(* Logix 5000 project; controller FV vendor 1 type 14 code 217 rev 31.11; software revision 31.00; part 5 of 63 *)
(* tags used below, declared in another part *)
   _1s_pulse : BOOL;
   FR_ALARM_RETURNED_STRING : STRING;
   FR_Crop_Event_Prefix : STRING;
   FR_Crop_Log_ID : DINT;
   FR_Event_Alarm_Tag : ALARM_DIGITAL;
   FR_Event_control_FIFO : CONTROL;
   FR_Event_control_FIFO_Operation_Type : CONTROL;
   FR_Event_Delay_For_Data : TIMER;
   FR_Event_Delay_For_PLC_Startup_Data : TIMER;
   FR_Event_Delay_Timer : TIMER;
   FR_Event_Delay_Timer_Off : TIMER;
   FR_Event_from_buffer : STRING;
   FR_Event_from_buffer_LogData1 : REAL;
   FR_Event_from_buffer_LogData2 : REAL;
   FR_Event_from_buffer_LogData3 : REAL;
   FR_Event_from_buffer_LogData4 : REAL;
   FR_Event_from_buffer_Operation_Type : DINT;
   FR_event_step : DINT;
   FR_Event_String_Last : STRING;
   FR_Event_Transact_Trigger_Tag : DINT;
   FR_Events_FIFO_Buffer : STRING[31];
   FR_Events_FIFO_Buffer_Operation_Type : DINT[31];
   FR_Filling_Event_Prefix : STRING;
   FR_Filling_Log_ID : DINT;
   FR_Filtrate_Event_Prefix : STRING;
   FR_Filtrate_Log_ID : DINT;
   FR_FVs26_31_Cropping_Event : STRING;
   FR_FVs26_31_Filling_Event : STRING;
   FR_FVs26_31_Filtrate_Event : STRING;
   FR_FVs26_31_Green_Beer_Event : STRING;
   FR_GreenBeer_Event_Prefix : STRING;
   FR_GreenBeer_Log_ID : DINT;
   FR_Last_LogData_For_Op : REAL[30,20];
   FR_N100 : INT[265];   // FV FILLING
   FR_N100_6_alarm : ALARM_DIGITAL;
   FR_N100_6_Alarm_Ready : BOOL;
   FR_N100_6_Delayed : DINT;
   FR_N100_6_Delayed_Timer : TIMER;
   FR_N100_6_Fault_Returned : STRING;
   FR_N100_6_SQL_Done : DINT;
   FR_N100_7_alarm : ALARM_DIGITAL;
   FR_N100_7_Alarm_Ready : BOOL;
   FR_N100_7_Delayed : DINT;
   FR_N100_7_Delayed_Timer : TIMER;
   FR_N100_7_Delayed_Timer2 : TIMER;
   FR_N100_7_Fault_Returned : STRING;
   FR_N100_7_SQL_Done : DINT;
   FR_N100_8_Delayed : DINT;
   FR_N100_8_Delayed_Timer : TIMER;
   FR_N110 : INT[265];   // GREEN BEER Green Beer Main
   FR_N110_6_alarm : ALARM_DIGITAL;
   FR_N110_6_Alarm_Ready : BOOL;
   FR_N110_6_Delayed : DINT;
   FR_N110_6_Delayed_Timer : TIMER;
   FR_N110_6_Fault_Returned : STRING;
   FR_N110_6_SQL_Done : DINT;
   FR_N110_7_alarm : ALARM_DIGITAL;
   FR_N110_7_Alarm_Ready : BOOL;
   FR_N110_7_Delayed : DINT;
   FR_N110_7_Delayed_Timer : TIMER;
   FR_N110_7_Delayed_Timer2 : TIMER;
   FR_N110_7_Fault_Returned : STRING;
   FR_N110_7_SQL_Done : DINT;
   FR_N110_8_Delayed : DINT;
   FR_N110_8_Delayed_Timer : TIMER;
   FR_N120 : INT[265];   // YEAST CROP Yeast Cropping Main
   FR_N120_6_alarm : ALARM_DIGITAL;
   FR_N120_6_Alarm_Ready : BOOL;
   FR_N120_6_Delayed : DINT;
   FR_N120_6_Delayed_Timer : TIMER;
   FR_N120_6_Fault_Returned : STRING;
   FR_N120_6_SQL_Done : DINT;
   FR_N120_7_alarm : ALARM_DIGITAL;
   FR_N120_7_Alarm_Ready : BOOL;
   FR_N120_7_Delayed : DINT;
   FR_N120_7_Delayed_Timer : TIMER;
   FR_N120_7_Delayed_Timer2 : TIMER;
   FR_N120_7_Fault_Returned : STRING;
   FR_N120_7_SQL_Done : DINT;
   FR_N120_8_Delayed : DINT;
   FR_N120_8_Delayed_Timer : TIMER;
   FR_N130 : INT[265];   // FILTRATE Filtrate Return
   FR_N130_6_alarm : ALARM_DIGITAL;
   FR_N130_6_Alarm_Ready : BOOL;
   FR_N130_6_Delayed : DINT;
   FR_N130_6_Delayed_Timer : TIMER;
   FR_N130_6_Fault_Returned : STRING;
   FR_N130_6_SQL_Done : DINT;
   FR_N130_7_alarm : ALARM_DIGITAL;
   FR_N130_7_Alarm_Ready : BOOL;
   FR_N130_7_Delayed : DINT;
   FR_N130_7_Delayed_Timer : TIMER;
   FR_N130_7_Delayed_Timer2 : TIMER;
   FR_N130_7_Fault_Returned : STRING;
   FR_N130_7_SQL_Done : DINT;
   FR_N130_8_Delayed : DINT;
   FR_N130_8_Delayed_Timer : TIMER;
   FtoF_raw_input : REAL;
   FV_B22 : INT[255];   // YSVFILL_FL YSV filling process flags
   FV_B32 : INT[255];   // PITCH_FLGS YSV pitching control flags
   FV_B42 : INT[255];   // YSVCIP_FLG
   FV_B52 : INT[255];   // WASTE_FLG
   FV_B62 : INT[255];   // RESEED FLG
   FV_B82 : INT[255];   // YSTFILL FL YST filling process flags
   FV_B86 : INT[255];   // YSTCIP FL YST CIP process flag s
   FV_N101 : INT[255];   // FV INT Fermentation control integer workspace
   FV_N139 : INT[255];   // YST1
   FV_N140 : INT[255];   // YST2
   FV_N141 : INT[255];   // YSV1 DATA
   FV_N142 : INT[255];   // YSV2 DATA
   FV_N143 : INT[255];   // YSV3 DATA
   FV_N144 : INT[255];   // YST1 DATA
   FV_N145 : INT[255];   // YST2 DATA
   FV_N20 : INT[255];   // YSVFILL<PC YSV Filling data fro m PC
   FV_N21 : INT[255];   // YSVFILL>PC YSV Filling process data to PC and contr ol regs
   FV_N30 : INT[255];   // PITCH<PC YSV Pitching data fr om PC
   FV_N31 : INT[255];   // PITCH>PC YSV Pitching data at o PC and control reg isters
   FV_N40 : INT[255];   // YSVCIP<PC
   FV_N41 : INT[255];   // YSVCIP>PC
   FV_N50 : INT[255];   // WASTE<PC
   FV_N51 : INT[255];   // WASTE>PC
   FV_N60 : INT[255];   // RESEED<PC
   FV_N61 : INT[255];   // RESEED>PC
   FV_N81 : INT[255];   // YSTFILL>PC YST filling process data to PC and contr ol regs.

        [5]   // YST filling routine alarm parameter #1
        [15]   // YST filling current YST data file pointer
        [16]   // YST filling command processor current step
   FV_N81_4_alarm : ALARM_DIGITAL;
   FV_N81_4_Alarm_Ready : BOOL;
   FV_N81_4_Delayed_Timer2 : TIMER := (PRE := 1000);
   FV_N81_4_Fault_Returned : STRING;
   FV_N81_4_SQL_Done : DINT := -1;
   FV_N84 : INT[255] := ([1] := -32768, [2] := -32768, [3] := -32768, [4] := -32768, [5] := -32768, [6] := -32768, [7] := -32768);   // YSTCIP<PC YST CIP data from PC
        [0].3   // Continue YST CIP
        [1]   // YST CIP selected YST
        [0].5   // End YST CIP
        [0].0   // Initiate YST CIP startup
        [0].15   // YST CIP cancel startup
        [0]   // YST CIP selected command
        [0].1   // Start YST CIP
        [0].4   // Abort YST CIP
        [0].2   // Stop YST CIP
   FV_N85 : INT[255] := ([0] := 1, [2] := 1, [16] := 1);   // YSTCIP>PC YST CIP process data to PC and control r egs.
        [2].3   // YST CIP continue available
        [4]   // YST CIP routine alarm register
        [9]   // YST CIP PC- displayed current step
        [1]   // YST CIP process current step
        [3]   // YST CIP process restart step
        [2].2   // YST CIP stop available
        [2].1   // YST CIP start available
        [2].4   // YST CIP abort available
        [14]   // YST CIP current YST attemperation file pointer
        [16]   // YST CIP command processor current step
        [15]   // YST CIP current YST data file pointer
        [2].0   // YST CIP initiate startup available
        [2].5   // YST CIP end available
        [0]   // YST CIP status (0:Unavailable; 1:Idle; 2:Running; 3:Stopped; 4:Faulted)
   FV_N85_4_alarm : ALARM_DIGITAL;
   FV_N85_4_Alarm_Ready : BOOL;
   FV_N85_4_Delayed_Timer2 : TIMER := (PRE := 1000);
   FV_N85_4_Fault_Returned : STRING;
   FV_N85_4_SQL_Done : DINT := -1;
   FV_N88 : INT[255] := ([1] := 99, [10] := 1, [20] := 1, [22] := 2, [23] := 10, [24] := 137, [28] := 5, [34] := 11826, [35] := 11828, [36] := 12593, [37] := 12590, [38] := 12338, [40] := -16384, [42] := 2, [43] := 10, [44] := 137, [48] := 23, [54] := 14641, [55] := 11826, [56] := 13873, [57] := 11832, [58] := 12338, [59] := 13102, [60] := 56);   // YSP COMMS Data transferred to/ from yeast press PLC
        [20].0   // Comms.to Yeast Press PLC failed flag
        [1]   // This PLC -> YSP PLC target tank no.
        [11].0   // YSP PLC -> This PLC YST1 high level probe
        [11].1   // YST PLC -> This PLC YST2 high level probe
        [10].0   // YSP PLC -> This PLC comms.handshake flag
        [0].0   // This PLC -> YSP PLC comms.handshake flag
   FV_PITCH_ACT : ALIAS FOR FV_B32[0].0;   // YSV Pitching Process Active
   FV_PITCH_AVAILABL_CMD : ALIAS FOR FV_N31[2];   // YSV Pitching Available Commands
   FV_PITCH_CUR_STEP : ALIAS FOR FV_N31[1];   // YSV Pitching Current Step
   FV_PITCH_DIALOG_AVAIL : ALIAS FOR FV_N31[2].0;   // PLC>PC YSV Pitching Startup Dialog Button Available
   FV_PITCH_PSCAN : ALIAS FOR FV_B32[0].2;   // YSV Pitching Postscan oneshot
   FV_PITCH_RES_STEP : ALIAS FOR FV_N31[3];   // YSV Pitching Restart Step
   FV_PITCH_RUN : ALIAS FOR FV_B32[0].1;   // YSVPitching Running
   FV_PITCH_SELECTED_CMD : ALIAS FOR FV_N30[0];   // YSV Pitching Selected Command
   FV_PITCH_START_SELECT : ALIAS FOR FV_N30[0].0;   // PC>PLC YSV Pitching Startup Dialog Buttlon Selected
   FV_PITCH_STATUS : ALIAS FOR FV_N31[0];   // YSV Pitching Status
   FV_PUMP1 : PlantItem := (CW := 2#0000_0000_0000_0000_0000_0000_1000_0001, CheckTime := 8, DriveBits := 1);   // PUMP1
   FV_PUMP1_RawOutput : ALIAS FOR Remote_IO:4:O.Data.13;   // FV_PUMP1 Coolant recirc.valve 1
   FV_PUMP2 : PlantItem := (CW := 2#0000_0000_0000_0000_0000_0000_1010_0001, CheckTime := 8, DriveBits := 1);   // PUMP2
   FV_PUMP2_RawOutput : ALIAS FOR Remote_IO:4:O.Data.14;   // FV_PUMP2 Coolant recirc.valve 2
   FV_PUMP3 : PlantItem := (CheckTime := 8);   // PUMP3
   FV_PUMP3_RawOutput : ALIAS FOR Remote_IO:4:O.Data.15;   // FV_PUMP3 Coolant recirc.valve 3
   FV_PV550_DPTR : ALIAS FOR FV_N101[8];   // Fermenting Room PV550 data file pointer
   FV_PX1 : PlantItem := (CW := 2#0000_0000_0000_0100_0000_0000_0000_0001, CheckTime := 12, DebounceTime := 4);   // PX1
   FV_PX1_RawInput : ALIAS FOR Remote_IO:6:I.Data.13;   // FV_PX1 Water flush proxy switch
   FV_PX2 : PlantItem := (CW := 2#0000_0000_0000_0000_0000_0000_0010_0000);   // PX2
   FV_PX2_RawInput : ALIAS FOR Remote_IO:6:I.Data.14;   // FV_PX2 CIP supply proxy switch
   FV_PX3 : PlantItem := (CW := 2#0000_0000_0000_0100_0000_0000_0010_0001);   // PX3
   FV_PX3_RawInput : ALIAS FOR Remote_IO:6:I.Data.15;   // FV_PX3 YSV1 to reseeding main proxy switch
   FV_R2V1 : PlantItem := (CW := 2#0000_0000_0000_0000_0000_0000_0001_0000, CheckTime := 15, CheckTimer := 15);   // R2V1
   FV_R2V1_ALARM : ALARM_DIGITAL;
   FV_R2V1_C : ALIAS FOR Remote_IO:7:I.Data.6;
   FV_R2V1_DR : ALIAS FOR Remote_IO:5:O.Data.10;
   FV_R2V1_O : ALIAS FOR Remote_IO:7:I.Data.2;
   FV_R2V2 : PlantItem := (CW := 2#0000_0000_0000_0000_0000_0000_1000_1011, CheckTime := 4, CheckTimer := 4, DriveBits := 4);   // R2V2
   FV_R2V2_ALARM : ALARM_DIGITAL;
   FV_R2V2_C : ALIAS FOR Remote_IO:7:I.Data.7;
   FV_R2V2_DR : ALIAS FOR Remote_IO:5:O.Data.11;
   FV_R2V2_O : ALIAS FOR Remote_IO:7:I.Data.3;
   FV_R6 : CONTROL[5] := ([1].LEN := 3, [2].LEN := 3, [2].UL := 1, [3].LEN := 3);
   FV_RESEED_ACT : ALIAS FOR FV_B62[0].0;   // YSV Reseeding Process Active
   FV_RESEED_AV1 : ALIAS FOR FV_B62[1];
   FV_RESEED_AV2 : ALIAS FOR FV_B62[2];
   FV_RESEED_AV3 : ALIAS FOR FV_B62[3];
   FV_RESEED_AV4 : ALIAS FOR FV_B62[4];
   FV_RESEED_AV5 : ALIAS FOR FV_B62[5];
   FV_RESEED_AVAILABL_CMD : ALIAS FOR FV_N61[2];   // YSV Reseeding Available Commands
   FV_RESEED_CUR_STEP : ALIAS FOR FV_N61[1];   // YSV Reseeding Current Step
   FV_RESEED_DIALOG_AVAIL : ALIAS FOR FV_N61[2].0;   // PLC>PC YSV Reseeding Startup Dialog Button Available
   FV_RESEED_END : ALIAS FOR FV_B62[0].8;   // YSV Reseeding End Process Selected
   FV_RESEED_PSCAN : ALIAS FOR FV_B62[0].2;   // YSV Reseeding Postscan oneshot
   FV_RESEED_RES_STEP : ALIAS FOR FV_N61[3];   // YSV Reseeding Restart Step
   FV_RESEED_RUN : ALIAS FOR FV_B62[0].1;   // YSV Reseeding Running
   FV_RESEED_SELECTED_CMD : ALIAS FOR FV_N60[0];   // YSV Reseeding Selected Command
   FV_RESEED_START_SELECT : ALIAS FOR FV_N60[0].0;   // PC>PLC YSV Reseeding Startup Dialog Buttlon Selected
   FV_RESEED_STATUS : ALIAS FOR FV_N61[0];   // YSV Reseeding Status
   FV_RSLN_CLEAN : ALIAS FOR FV_B62[1].0;   // Reseeding line clean flag
   FV_SFile : INT[255] := ([4] := 19904, [13] := 3, [37] := 2020, [38] := 7, [39] := 31, [40] := 13, [41] := 9, [42] := 50);   // SLC Equivalent System File, So Original Code Can Remain
        [1].15   // First Scan Flag
        [37]   // Clock Calendar Year
        [41]   // Clock Calendar Minutes
        [53]   // Calendar Day 1 = Monday
        [40]   // Clock Calendar Hours
        [42]   // Clock Calendar Minute
   FV_SOV1 : PlantItem := (CheckTime := 8);   // SOV1
   FV_SOV1_RawOutput : ALIAS FOR Remote_IO:5:O.Data.6;   // FV_SOV1 Air supply to reseed pump
   FV_SOV2 : PlantItem := (CheckTime := 8);   // SOV2
   FV_SOV2_RawOutput : ALIAS FOR Remote_IO:5:O.Data.7;   // FV_SOV2 Air supply to reseed pump
   FV_T102 : TIMER[20] := ([0].PRE := 360000, [0].ACC := 298181, [0].EN := 1, [0].TT := 1);
   FV_T16 : TIMER[10] := ([0].PRE := 8000, [0].ACC := 3002, [0].EN := 1, [0].TT := 1);
   FV_T212 : TIMER[5] := ([0].PRE := 3000, [0].EN := 1, [0].DN := 1, [1].PRE := 3000, [1].EN := 1, [1].DN := 1, [2].PRE := 3000, [2].ACC := 3000);
   FV_T23 : TIMER[10] := ([0].PRE := 300000);
   FV_T33 : TIMER[10] := ([0].PRE := 300000, [1].PRE := 60000, [2].PRE := 10000);
   FV_T4 : TIMER[10] := ([0].PRE := 2000, [1].PRE := 300000, [2].PRE := 2500, [2].ACC := 50, [2].EN := 1, [2].TT := 1, [3].PRE := 300000, [3].ACC := 300001, [3].EN := 1, [3].DN := 1, [4].PRE := 3300000, [4].ACC := 2309456, [4].EN := 1, [4].TT := 1, [5].PRE := 3600000, [6].PRE := 60000, [8].PRE := 10000, [9].PRE := 10000);
   FV_T43 : TIMER[10] := ([0].PRE := 300000);
   FV_T53 : TIMER[10] := ([0].PRE := 300000, [2].PRE := 10000);
   FV_T63 : TIMER[20] := ([0].PRE := 60000, [3].PRE := 120000, [3].ACC := 82385, [4].PRE := 13000, [5].PRE := 16000, [6].PRE := 30000, [7].PRE := 4000, [8].PRE := 4000);
   FV_T73 : TIMER[10] := ([0].PRE := 300000, [1].PRE := 30000, [2].PRE := 20000);
   FV_T83 : TIMER[5] := ([0].PRE := 300000);
   FV_T87 : TIMER[2] := ([0].PRE := 300000);
   FV_T89 : TIMER[5] := ([0].PRE := 3000, [0].ACC := 1745, [0].EN := 1, [0].TT := 1, [1].PRE := 10000, [2].PRE := 10000, [2].ACC := 10001, [2].EN := 1, [2].DN := 1);
   FV_to_data_file : DINT;
   FV_to_data_offset : DINT;
   FV_TTX_YS_001_AI : PlantItem := (CW := 2#0000_0000_0000_0000_1100_0000_0000_0000, CheckTime := 10, CheckTimer := 10, Scaled := 18.41875, RawInput := 6947.0);   // TTX_YS_001
   FV_TTX_YS_001_AI_RawInput : ALIAS FOR Remote_IO:8:I.Ch00Data;   // Real Analog Input , Do Not Use In Code
   FV_TTX_YS_002_AI : PlantItem := (CW := 2#0000_0000_0000_0000_1000_0000_0000_0000, CheckTime := 10, CheckTimer := 10, Scaled := 9.6625, RawInput := 5546.0);   // TTX_YS_002
   FV_TTX_YS_002_AI_RawInput : ALIAS FOR Remote_IO:8:I.Ch01Data;   // Real Analog Input , Do Not Use In Code
   FV_value_to_set : INT;
   FV_WASTE_ACT : ALIAS FOR FV_B52[0].0;   // YSV To Waste Process Active
   FV_WASTE_AVAILABL_CMD : ALIAS FOR FV_N51[2];   // YSV To Waste Available Commands
   FV_WASTE_CUR_STEP : ALIAS FOR FV_N51[1];   // YSV To Waste Current Step
   FV_WASTE_DIALOG_AVAIL : ALIAS FOR FV_N51[2].0;   // PLC>PC YSV To Waste Startup Dialog Button Available
   FV_WASTE_PSCAN : ALIAS FOR FV_B52[0].2;   // YSV To Waste Postscan oneshot
   FV_WASTE_RES_STEP : ALIAS FOR FV_N51[3];   // YSV To Waste Restart Step
   FV_WASTE_RUN : ALIAS FOR FV_B52[0].1;   // YSV To Waste Running
   FV_WASTE_SELECTED_CMD : ALIAS FOR FV_N50[0];   // YSV To Waste Selected Command
   FV_WASTE_START_SELECT : ALIAS FOR FV_N50[0].0;   // PC>PLC YSV To Waste Startup Dialog Buttlon Selected
   FV_WASTE_STATUS : ALIAS FOR FV_N51[0];   // YSV To Waste Status
   FV_word_offset : INT;
   FV_WYT1R : PlantItem := (CW := 2#0000_0000_0000_0000_0000_1100_0000_0000, CheckTime := 8, CheckTimer := 8);   // WYT1R
   FV_WYT1R_ALARM : ALARM_DIGITAL;
   FV_WYT1R_D : ALIAS FOR Remote_IO:5:O.Data.14;
   FV_WYT1R_R : ALIAS FOR Remote_IO:7:I.Data.20;
   FV_WYT2R : PlantItem := (CW := 2#0000_0000_0000_0000_0000_1100_1000_1011, CheckTime := 8, CheckTimer := 8, DriveBits := 1);   // WYT2R
   FV_WYT2R_ALARM : ALARM_DIGITAL;
   FV_WYT2R_D : ALIAS FOR Remote_IO:5:O.Data.15;
   FV_WYT2R_R : ALIAS FOR Remote_IO:7:I.Data.21;
   FV_WYTR1 : PlantItem := (CW := 2#0000_0000_0000_0000_0000_0000_0001_0000, CheckTime := 10, CheckTimer := 10);   // WYTR1
   FV_WYTR1_ALARM : ALARM_DIGITAL;
   FV_WYTR1_C : ALIAS FOR Remote_IO:7:I.Data.4;
   FV_WYTR1_DR : ALIAS FOR Remote_IO:5:O.Data.8;
   FV_WYTR1_O : ALIAS FOR Remote_IO:7:I.Data.0;
   FV_WYTR2 : PlantItem := (CW := 2#0000_0000_0000_0000_0000_0000_0001_0000, CheckTime := 4, CheckTimer := 4);   // WYTR2
   FV_WYTR2_ALARM : ALARM_DIGITAL;
   FV_WYTR2_C : ALIAS FOR Remote_IO:7:I.Data.5;
   FV_WYTR2_DR : ALIAS FOR Remote_IO:5:O.Data.9;
   FV_WYTR2_O : ALIAS FOR Remote_IO:7:I.Data.1;
   FV_Yeast_Press_Blunger_Comms : MESSAGE;
        MessageParameters(ServiceCode := 16#0fa2, LocalElement := FV_N88[10], ...)
   FV_YSPC_FAIL : ALIAS FOR FV_N88[20].0;   // Comms.to Yeast Press PLC failed flag
   FV_YST01_LTX501_Fill_Lvl_OK : TIMER := (PRE := 1000);
   FV_YST02_LTX501_Fill_Lvl_OK : TIMER := (PRE := 1000);
   FV_YST1_FV : ALIAS FOR FV_N139[0];   // YST1 attemperation control data
   FV_YST1_HL_SP : DINT := 145;
   FV_YST1_STATUS : ALIAS FOR FV_N144[0];   // YST1 current operation
   FV_YST2_FV : ALIAS FOR FV_N140[0];   // YST2 attemperation control data
   FV_YST2_HL_SP : DINT := 145;
   FV_YST2_STATUS : ALIAS FOR FV_N145[0];   // YST2 current operation
   FV_YSTCIP_ACT : ALIAS FOR FV_B86[0].0;   // YST CIP process active
   FV_YSTCIP_Log_ID : DINT := 10;
   FV_YSTCIP_RESTART : ALIAS FOR FV_N85[3];   // YST CIP process restart step
   FV_YSTCIP_RUN : ALIAS FOR FV_B86[0].1;   // YST CIP running
   FV_YSTCIP_STATUS : ALIAS FOR FV_N85[0];   // YST CIP status (0:Unavailable; 1:Idle; 2:Running; 3:Stopped; 4:Faulted)
   FV_YSTCIP_STEP : ALIAS FOR FV_N85[1];   // YST CIP process current step
   FV_YSTFILL_ACT : ALIAS FOR FV_B82[0].0;   // YST filling process active
   FV_YSTFILL_Log_ID : DINT := 3;
   FV_YSTFILL_PSCAN : ALIAS FOR FV_B82[0].2;   // YST filling postscan oneshot
   FV_YSTFILL_RESTART : ALIAS FOR FV_N81[3];   // YST filling restart step
   FV_YSTFILL_RUN : ALIAS FOR FV_B82[0].1;   // YST filling process running
   FV_YSTFILL_STATUS : ALIAS FOR FV_N81[0];   // YST filling status (0:Unavailable; 1:Idle; 2:Running; 3:Stopped; 4:Faulted)
   FV_YSTFILL_STEP : ALIAS FOR FV_N81[1];   // YST filling current step
   FV_YSTs_CIP_Vessel_Event : STRING;
   FV_YSTs_CIP_Vessel_Event_Prefix : STRING := 'YST 1 ';
   FV_YSTs_Filling_Event : STRING;
   FV_YSTs_Filling_Event_Prefix : STRING := 'YST 1 ';
   FV_YSV1_RSR_MODE : ALIAS FOR FV_N141[3];   // YSV1 Rouser Mode 0=Auto 1 = Manual On 2 = Manual Off
   FV_YSV1_STATUS : ALIAS FOR FV_N141[0];   // YSV1 Current Operation
   FV_YSV1_TTX01_AI : PlantItem := (CW := 2#0000_0000_0000_0000_1000_0000_0000_0000, CheckTime := 10, CheckTimer := 10, Scaled := 4.640625, RawInput := 8685.0);   // YSV1_TTX01
   FV_YSV1_TTX01_AI_RawInput : ALIAS FOR Remote_IO:13:I.Ch1Data;   // Real Analog Input , Do Not Use In Code
   FV_YSV1_WEIGHT : ALIAS FOR FV_N141[2];   // YSV1 current weight kg*10
   FV_YSV1_WTX01_AI : PlantItem := (CW := 2#0000_0000_0000_0000_1000_0000_0000_0000, CheckTime := 10, CheckTimer := 10, Scaled := 51.7575, RawInput := 5648.0);   // YSV1_WTX01
   FV_YSV1_WTX01_AI_RawInput : ALIAS FOR Remote_IO:13:I.Ch6Data;   // Real Analog Input , Do Not Use In Code
   FV_YSV1CV : PlantItem := (CW := 2#0000_0000_0000_0000_0000_0000_0100_0000, CheckTime := 8);   // YSV1CV
   FV_YSV1CV_RawOutput : ALIAS FOR Remote_IO:5:O.Data.12;   // FV_YSV1CV
   FV_YSV1J : PlantItem := (CW := 2#0000_0000_0000_0000_0000_0000_1000_0001, CheckTime := 8, DriveBits := 1);   // YSV1J
   FV_YSV1J_RawOutput : ALIAS FOR Remote_IO:4:O.Data.9;   // FV_YSV1J YSV 1 cooling valve
   FV_YSV1R : PlantItem := (CW := 2#0000_0000_0000_0000_0000_1100_0000_0000, CheckTime := 8, CheckTimer := 8);   // YSV1R
   FV_YSV1R_ALARM : ALARM_DIGITAL;
   FV_YSV1R_D : ALIAS FOR Remote_IO:4:O.Data.10;   // YSV 1 rouser
   FV_YSV1R_R : ALIAS FOR Remote_IO:6:I.Data.12;   // YSV 1 Rouser running f/b
   FV_YSV2_STATUS : ALIAS FOR FV_N142[0];   // YSV2 Current Operation
   FV_YSV2_TTX01_AI : PlantItem := (CW := 2#0000_0000_0000_0000_1000_0000_0000_0000, CheckTime := 10, CheckTimer := 10, Scaled := 3.1531248, RawInput := 8209.0);   // YSV2_TTX01
   FV_YSV2_TTX01_AI_RawInput : ALIAS FOR Remote_IO:13:I.Ch2Data;   // Real Analog Input , Do Not Use In Code
   FV_YSV2_WEIGHT : ALIAS FOR FV_N142[2];   // YSV2 current weight kg*10
   FV_YSV2_WTX01_AI : PlantItem := (CW := 2#0000_0000_0000_0000_1000_0000_0000_0000, CheckTime := 10, CheckTimer := 10, Scaled := 155.11562, RawInput := 11091.0);   // YSV2_WTX01
   FV_YSV2_WTX01_AI_RawInput : ALIAS FOR Remote_IO:13:I.Ch5Data;   // Real Analog Input , Do Not Use In Code
   FV_YSV2CV : PlantItem := (CW := 2#0000_0000_0000_0000_0000_0000_1000_0001, CheckTime := 8, DriveBits := 1);   // YSV2CV
   FV_YSV2CV_RawOutput : ALIAS FOR Remote_IO:5:O.Data.13;   // FV_YSV2CV
   FV_YSV2J : PlantItem := (CW := 2#0000_0000_0000_0000_0000_0000_1000_0001, CheckTime := 8, DriveBits := 1);   // YSV2J
   FV_YSV2J_RawOutput : ALIAS FOR Remote_IO:4:O.Data.11;   // FV_YSV2J YSV 2 cooling valve
   FV_YSV2O : PlantItem := (CheckTime := 8);   // YSV2O
   FV_YSV2O_RawOutput : ALIAS FOR Remote_IO:4:O.Data.4;   // FV_YSV2O YSV 2 outlet valve
   FV_YSV2R : PlantItem := (CheckTime := 8);   // YSV2R
   FV_YSV2R_RawOutput : ALIAS FOR Remote_IO:4:O.Data.12;   // FV_YSV2R YSV 2 rouser
   FV_YSV3_STATUS : ALIAS FOR FV_N143[0];   // YSV3 Current Operation
   FV_YSV3_TTX01_AI : PlantItem := (CW := 2#0000_0000_0000_0000_1000_0000_0000_0000, CheckTime := 10, CheckTimer := 10, Scaled := 21.153126, RawInput := 13969.0);   // YSV3_TTX01
   FV_YSV3_TTX01_AI_RawInput : ALIAS FOR Remote_IO:13:I.Ch3Data;   // Real Analog Input , Do Not Use In Code
   FV_YSV3_WEIGHT : ALIAS FOR FV_N143[2];   // YSV3 current weight kg*10
   FV_YSV3_WTX01_AI : PlantItem := (CW := 2#0000_0000_0000_0000_1000_0000_0000_0000, CheckTime := 10, CheckTimer := 10, Scaled := 0.0625, RawInput := 4002.0);   // YSV3_WTX01
   FV_YSV3_WTX01_AI_RawInput : ALIAS FOR Remote_IO:13:I.Ch4Data;   // Real Analog Input , Do Not Use In Code
   FV_YSV3J : PlantItem := (CheckTime := 8);   // YSV3J
   FV_YSV3J_RawOutput : ALIAS FOR Remote_IO:4:O.Data.7;   // FV_YSV3J YSV 3 cooling valve
   FV_YSV3O : PlantItem := (CheckTime := 8);   // YSV3O
   FV_YSV3O_RawOutput : ALIAS FOR Remote_IO:4:O.Data.6;   // FV_YSV3O YSV 3 outlet valve
   FV_YSV3R : PlantItem := (CheckTime := 8);   // YSV3R
   FV_YSV3R_RawOutput : ALIAS FOR Remote_IO:4:O.Data.8;   // FV_YSV3R YSV 3 rouser
   FV_YSVCIP_ACT : ALIAS FOR FV_B42[0].0;   // YSV CIP Process Active
   FV_YSVCIP_AVAILABL_CMD : ALIAS FOR FV_N41[2];   // YSV CIP Available Commands
   FV_YSVCIP_CUR_STEP : ALIAS FOR FV_N41[1];   // YSV CIP Current Step
   FV_YSVCIP_DIALOG_AVAIL : ALIAS FOR FV_N41[2].0;   // PLC>PC YSV CIP Startup Dialog Button Available
   FV_YSVCIP_END : ALIAS FOR FV_B42[0].8;   // YSV CIP End Process Selected
   FV_YSVCIP_PSCAN : ALIAS FOR FV_B42[0].2;   // YSV CIP Postscan oneshot
   FV_YSVCIP_RES_STEP : ALIAS FOR FV_N41[3];   // YSV CIP Restart Step
   FV_YSVCIP_RUN : ALIAS FOR FV_B42[0].1;   // YSV CIP Running
   FV_YSVCIP_SELECTED_CMD : ALIAS FOR FV_N40[0];   // YSV CIP Selected Command
   FV_YSVCIP_START_SELECT : ALIAS FOR FV_N40[0].0;   // PC>PLC YSV CIP Startup Dialog Buttlon Selected
   FV_YSVCIP_STATUS : ALIAS FOR FV_N41[0];   // YSV CIP Status
   FV_YSVCIPLINE_Log_ID : DINT := 7;
   FV_YSVCIPVESSEL_Log_ID : DINT := 6;
   FV_YSVFILL_ACT : ALIAS FOR FV_B22[0].0;   // YSV Filling Process Active
   FV_YSVFILL_AVAILABL_CMD : ALIAS FOR FV_N21[2];   // YSV Filling Available Commands
   FV_YSVFILL_CUR_STEP : ALIAS FOR FV_N21[1];   // YSV Filling Current Step
   FV_YSVFILL_DIALOG_AVAIL : ALIAS FOR FV_N21[2].0;   // PLC>PC YSV Filling Startup Dialog Button Available
   FV_YSVFILL_END : ALIAS FOR FV_B22[0].8;   // YSV Filling End Process Selected
   FV_YSVFILL_Log_ID : DINT := 4;
   FV_YSVFILL_PSCAN : ALIAS FOR FV_B22[0].2;   // YSV Filling Postscan oneshot
   FV_YSVFILL_RES_STEP : ALIAS FOR FV_N21[3];   // YSV Filling Restart Step
   FV_YSVFILL_RUN : ALIAS FOR FV_B22[0].1;   // YSV Filling Running
   FV_YSVFILL_SELECTED_CMD : ALIAS FOR FV_N20[0];   // YSV Filling Selected Command
   FV_YSVFILL_START_SELECT : ALIAS FOR FV_N20[0].0;   // PC>PLC YSV Filling Startup Dialog Buttlon Selected
   FV_YSVFILL_STATUS : ALIAS FOR FV_N21[0];   // YSV Filling Status
   FV_YSVPITCH_Log_ID : DINT := 5;
   FV_YSVPitching_AmountAtEnd : REAL := 155.68437;
   FV_YSVRESEED_Log_ID : DINT := 9;
   FV_YSVs_CIP_Line_Event : STRING;
   FV_YSVs_CIP_Line_Event_prefix : STRING;
   FV_YSVs_CIP_vessel_Event : STRING;
   FV_YSVs_CIP_vessel_Event_Prefix : STRING := 'YSV 2 ';
   FV_YSVs_Filling_Event : STRING;
   FV_YSVs_Filling_Event_Prefix : STRING := 'YSV 2 ';
   FV_YSVs_Pitching_Event : STRING;
   FV_YSVs_Pitching_Event_Prefix : STRING := 'YSV 2 ';
   FV_YSVs_reseeding_event : STRING;
   FV_YSVs_reseeding_event_prefix : STRING := 'YSV 1 ';
   FV_YSVs_to_waste_event : STRING;
   FV_YSVs_to_waste_event_prefix : STRING := 'YSV 2 ';
   FV_YSVTOWASTE_Log_ID : DINT := 8;
   FV_YSVWaste_AmountAtEnd : REAL := 0.56874996;
   go_test_operation_temp : BOOL;
   indirect_bit_temp : INT := 7;
   Item_Faults_Are_Latched : BOOL;
   Item_Simulation_Flag : BOOL;
   ItoF_raw_input : INT := 5648;
   Mike_141019 : BOOL := 1;
   MV_Read_YST : MESSAGE;
        MessageParameters(ServiceCode := 16#004c, LocalElement := MV_YST_Levels[0], ...)
   MV_Read_YST_TMR : TIMER := (PRE := 500, ACC := 485, EN := 1, TT := 1);
   MV_YST_Levels : REAL[2] := ([0] := 0.028125001, [1] := 79.640625);
        [0]   // YST1 Level
        [1]   // YST2 Level
   One_Minute_One_Scan : BOOL;
   One_Minute_One_Scan_Timer : TIMER := (PRE := 60000, ACC := 51773, EN := 1, TT := 1);
   One_Second_1_scan : BOOL;
   One_Second_One_Scan : ALIAS FOR One_Second_1_scan;
   One_Second_Toggle : BOOL := 1;
   overrange_RIO_analog_value : REAL;
   Pitching_transaction_locked_timer : TIMER := (PRE := 10000);
   Pitching_transaction_log : DINT;
   Pitching_transaction_log_delay : DINT;
   Pitching_transaction_log_Done : DINT := -1;
   Pitching_transaction_log_timer : TIMER := (PRE := 10000);
   rack_simulation_flag : BOOL;
   Reseeding_transaction_locked_timer : TIMER := (PRE := 10000);
   Reseeding_transaction_log : DINT;
   Reseeding_transaction_log_delay : DINT;
   Reseeding_transaction_log_Done : DINT := -1;
   Reseeding_transaction_log_timer : TIMER := (PRE := 10000);
   reset_msg_interval : BOOL;
   Scada_Pump_Fault_No : DINT := 20001;
   Scada_Pump_H_Fault_No : DINT;
   Scada_Pump_T_Fault_No : DINT;
   Scada_Valve_Fault_No : DINT := 10001;
   scada_watchdog : DINT := 15;
   scada_watchdog_tmr : TIMER := (PRE := 1000);
   scada_watchdog_tmr_off : TIMER := (PRE := 1000, ACC := 242, EN := 1, TT := 1);
   scale_analog_int : DINT := 12000;
   scale_analog_result : REAL := 1142.0016;
   scale_eu_max : REAL := 502.5;
   scale_eu_max_int : DINT := 300;
   scale_eu_min : REAL;
   scale_eu_min_int : DINT := 200;
   scale_raw_input : REAL := 11091.0;
   scale_raw_max : REAL := 20000.0;
   scale_raw_max_int : DINT := 120;
   scale_raw_min : REAL := 4000.0;
   scale_raw_min_int : DINT;
   scale_routine_active : BOOL := 1;
   scale_temp : REAL := 0.03140625;
   TempChecktime : DINT := 32;
   template_analog_input : PlantItem;
   template_analog_input_RawInput : REAL;
   template_analog_output : PlantItem;
   template_analog_output_RawOutput : REAL;
   template_boolean : BOOL;
   template_input : PlantItem;
   template_input_RawInput : ALIAS FOR template_boolean;
   template_output : PlantItem;
   template_output_RawOutput : ALIAS FOR template_boolean;   // P04CHILLRUN Chiller Run Signal
   template_pump : PlantItem;
   template_pump_D : ALIAS FOR template_boolean;   // auto start vacuum pump 1
   template_pump_H : ALIAS FOR template_boolean;   // vacuum pump 1 auto avail
   template_pump_ISOL : ALIAS FOR template_boolean;
   template_pump_R : ALIAS FOR template_boolean;   // vacuum pump 1 running
   template_valve : PlantItem;
   template_valve_C : ALIAS FOR template_boolean;   // skim manifold to ycv2 drain valve closed
   template_valve_DR : ALIAS FOR template_boolean;   // drive open skim manifold to ycv2 drain valve
   template_valve_O : ALIAS FOR template_boolean;   // skim manifold to ycv2 drain valve opened
   tempv : DINT;
   Test_Cropping_done : BOOL := 1;
   underrange_RIO_analog_value : REAL;
   Unused_Healthy_Feedback : BOOL := 1;
   Unused_NotTripped_Feedback : BOOL := 1;
   YP_ALARM_ACCEPT : ALIAS FOR YP_B103[1].2;
   YP_ALARM_ACCEPT_OS_FLAG : ALIAS FOR YP_B103[1].0;
   YP_AV1 : PlantItem := (CW := 2#0000_0000_0000_0000_0000_0000_0001_0000, CheckTime := 15, CheckTimer := 15);   // AV1
   YP_AV10_MANUAL : ALIAS FOR YP_N50[9];
   YP_AV10_REQUIRED : ALIAS FOR YP_B30[0].14;   // BLUNGER TRANSFER PUMP
   YP_AV1_ALARM : ALARM_DIGITAL;
   YP_AV1_CLOSE_FAULT : ALIAS FOR YP_B92[0].1;
   YP_AV1_CLOSE_FLT_TIMER : ALIAS FOR YP_T20[1];
   YP_AV1_DR : ALIAS FOR RIO_Rack_3:3:O.Data.3;
   YP_AV1_MANUAL : ALIAS FOR YP_N50[0];
   YP_AV1_O : ALIAS FOR RIO_Rack_3:1:I.Data.0;
   YP_AV1_OPEN_FAULT : ALIAS FOR YP_B92[0].0;
   YP_AV1_OPEN_FLT_TIMER : ALIAS FOR YP_T20[0];
   YP_AV1_REQUIRED : ALIAS FOR YP_B30[0].3;
   YP_AV2 : PlantItem := (CW := 2#0000_0000_0000_0000_0000_0001_0001_0000, CheckTime := 15, CheckTimer := 15);   // AV2
   YP_AV2_ALARM : ALARM_DIGITAL;
   YP_AV2_CLOSE_FAULT : ALIAS FOR YP_B92[0].3;
   YP_AV2_CLOSE_FLT_TIMER : ALIAS FOR YP_T20[3];
   YP_AV2_DR : ALIAS FOR RIO_Rack_3:3:O.Data.5;
   YP_AV2_MANUAL : ALIAS FOR YP_N50[1];
   YP_AV2_O : ALIAS FOR RIO_Rack_3:1:I.Data.2;
   YP_AV2_OPEN_FAULT : ALIAS FOR YP_B92[0].2;
   YP_AV2_OPEN_FLAG : ALIAS FOR YP_B3[0].2;
   YP_AV2_OPEN_FLT_TIMER : ALIAS FOR YP_T20[2];
   YP_AV2_REQUIRED : ALIAS FOR YP_B30[0].5;
   YP_AV3 : PlantItem := (CW := 2#0000_0000_0000_0000_0000_0000_0001_0000, CheckTime := 15, CheckTimer := 15);   // AV3
   YP_AV3_ALARM : ALARM_DIGITAL;
   YP_AV3_CLOSE_FAULT : ALIAS FOR YP_B92[0].5;
   YP_AV3_CLOSE_FLT_TIMER : ALIAS FOR YP_T20[5];
   YP_AV3_DR : ALIAS FOR RIO_Rack_3:3:O.Data.6;
   YP_AV3_MANUAL : ALIAS FOR YP_N50[2];
   YP_AV3_O : ALIAS FOR RIO_Rack_3:1:I.Data.4;
   YP_AV3_OPEN_FAULT : ALIAS FOR YP_B92[0].4;
   YP_AV3_OPEN_FLAG : ALIAS FOR YP_B3[0].4;
   YP_AV3_OPEN_FLT_TIMER : ALIAS FOR YP_T20[4];
   YP_AV3_REQUIRED : ALIAS FOR YP_B30[0].6;
   YP_AV4 : PlantItem := (CW := 2#0000_0000_0000_0000_0000_0000_0001_0000, CheckTime := 15, CheckTimer := 15);   // AV4
   YP_AV4_ALARM : ALARM_DIGITAL;
   YP_AV4_CLOSE_FAULT : ALIAS FOR YP_B92[0].7;
   YP_AV4_CLOSE_FLT_TIMER : ALIAS FOR YP_T20[7];
   YP_AV4_DR : ALIAS FOR RIO_Rack_3:3:O.Data.7;
   YP_AV4_MANUAL : ALIAS FOR YP_N50[3];
   YP_AV4_O : ALIAS FOR RIO_Rack_3:1:I.Data.6;
   YP_AV4_OPEN_FAULT : ALIAS FOR YP_B92[0].6;
   YP_AV4_OPEN_FLAG : ALIAS FOR YP_B3[0].6;
   YP_AV4_OPEN_FLT_TIMER : ALIAS FOR YP_T20[6];
   YP_AV4_REQUIRED : ALIAS FOR YP_B30[0].7;
   YP_AV5 : PlantItem := (CW := 2#0000_0000_0000_0000_0000_0000_0001_0000, CheckTime := 15, CheckTimer := 15);   // AV5
   YP_AV5_ALARM : ALARM_DIGITAL;
   YP_AV5_CLOSE_FLT_TIMER : ALIAS FOR YP_T20[9];
   YP_AV5_CLSOE_FAULT : ALIAS FOR YP_B92[0].9;
   YP_AV5_DR : ALIAS FOR RIO_Rack_3:3:O.Data.8;
   YP_AV5_O : ALIAS FOR RIO_Rack_3:1:I.Data.8;
   YP_AV5_OPEN_FAULT : ALIAS FOR YP_B92[0].8;
   YP_AV5_OPEN_FLAG : ALIAS FOR YP_B3[0].8;
   YP_AV5_OPEN_FLT_TIMER : ALIAS FOR YP_T20[8];
   YP_AV5_REQUIRED : ALIAS FOR YP_B30[0].8;
   YP_AV6 : PlantItem := (CW := 2#0000_0000_0000_0000_0000_0000_0001_0000, CheckTime := 15, CheckTimer := 15);   // AV6
   YP_AV6_ALARM : ALARM_DIGITAL;
   YP_AV6_CLOSE_FAULT : ALIAS FOR YP_B92[0].11;
   YP_AV6_CLOSE_FLT_TIMER : ALIAS FOR YP_T20[11];
   YP_AV6_DR : ALIAS FOR RIO_Rack_3:3:O.Data.9;
   YP_AV6_MANUAL : ALIAS FOR YP_N50[5];
   YP_AV6_O : ALIAS FOR RIO_Rack_3:1:I.Data.10;
   YP_AV6_OPEN_FAULT : ALIAS FOR YP_B92[0].10;
   YP_AV6_OPEN_FLAG : ALIAS FOR YP_B3[0].10;
   YP_AV6_OPEN_FLT_TIMER : ALIAS FOR YP_T20[10];
   YP_AV6_RQUIRED : ALIAS FOR YP_B30[0].9;
   YP_AV7 : PlantItem := (CW := 2#0000_0000_0000_0000_0000_0000_0001_0000, CheckTime := 15, CheckTimer := 15);   // AV7
   YP_AV7_ALARM : ALARM_DIGITAL;
   YP_AV7_CLOSE_FAULT : ALIAS FOR YP_B92[0].13;
   YP_AV7_CLOSE_FLT_TIMER : ALIAS FOR YP_T20[13];
   YP_AV7_DR : ALIAS FOR RIO_Rack_3:3:O.Data.10;
   YP_AV7_MANUAL : ALIAS FOR YP_N50[6];
   YP_AV7_O : ALIAS FOR RIO_Rack_3:1:I.Data.12;
   YP_AV7_OPEN_FAULT : ALIAS FOR YP_B92[0].12;
   YP_AV7_OPEN_FLAG : ALIAS FOR YP_B3[0].12;
   YP_AV7_OPEN_FLT_TIMER : ALIAS FOR YP_T20[12];
   YP_AV7_REQUIRED : ALIAS FOR YP_B30[0].10;
   YP_AV8 : PlantItem := (CW := 2#0000_0000_0000_0000_0000_0000_0001_0000, CheckTime := 15, CheckTimer := 15);   // AV8
   YP_AV8_ALARM : ALARM_DIGITAL;
   YP_AV8_CLOSE_FAULT : ALIAS FOR YP_B92[0].15;
   YP_AV8_CLOSE_FLT_TIMER : ALIAS FOR YP_T20[15];
   YP_AV8_DR : ALIAS FOR RIO_Rack_3:3:O.Data.11;
   YP_AV8_MANUAL : ALIAS FOR YP_N50[7];
   YP_AV8_O : ALIAS FOR RIO_Rack_3:1:I.Data.14;
   YP_AV8_OPEN_FAULT : ALIAS FOR YP_B92[0].14;
   YP_AV8_OPEN_FLAG : ALIAS FOR YP_B3[0].14;
   YP_AV8_OPEN_FLT_TIMER : ALIAS FOR YP_T20[14];
   YP_AV8_REQUIRED : ALIAS FOR YP_B30[0].11;
   YP_AV9_MANUAL : ALIAS FOR YP_N50[8];
   YP_B103 : INT[15] := ([0] := 1);   // Original N File From SLC, No Description Available
        [0].0   // Yeast Press CIP Heartbeat Fault
        [2].2   // Channel 1 CIP Active
        [2].3   // Channel 2 CIP Active
        [3].0   // START BLUNGER WATER FILL FROM PV
        [3].1   // STOP BLUNGER WATER FILL FROM PV
        [4].0   // Fill Cycle Controls Force End Of Cycle
   YP_B103_1_1_Storagebit : BOOL;
   YP_B3 : INT[7] := ([1] := 4);   // BINARY
        [1].1   // Press closed
        [1].2   // Press open microswitch should trigger start conveyor
   YP_B30 : INT[37];   // Original N File From SLC, No Description Available
        [0].14   // BLUNGER TRANSFER PUMP
   YP_B31 : INT[37] := ([31] := 16);   // Original N File From SLC, No Description Available
   YP_B92 : INT[105] := ([2] := 4, [20] := 2, [22] := 4, [60] := 2, [62] := 4);   // Original N File From SLC, No Description Available
   YP_BEAT_FROM_FV : ALIAS FOR YP_N10[10].0;
   YP_BEAT_TO_FV_PLC : ALIAS FOR YP_N10[0].0;
   YP_BLUNG_OV : PlantItem;   // BLUNG_OV
   YP_BLUNG_OV_RawInput : ALIAS FOR RIO_Rack_3:2:I.Data.1;   // YP_BLUNG_OV
   YP_BLUNGER_DRAIN_IDLE : ALIAS FOR YP_N40[3].0;   // BLUNGER DRAIN/RANSFER TO YST IDLE FLAG
   YP_BLUNGER_DRAIN_TIMER : ALIAS FOR YP_T21[2];
   YP_BLUNGER_FILL_SP_1 : ALIAS FOR YP_N55[32];   // Blunger Water Feed Feed Timer 1
   YP_BLUNGER_FILL_TIMER : ALIAS FOR YP_N55[31];   // BLUNGER FILL TIMER SELECTED FROM PV
   YP_BLUNGER_FILL_TIMER_2 : ALIAS FOR YP_N55[33];   // Blunger Water Feed Feed Timer 2
   YP_BLUNGER_FILL_TIMER_3 : ALIAS FOR YP_N55[34];   // Blunger Water Feed Feed Timer 3
   YP_BLUNGER_TRANS_DEST : ALIAS FOR YP_N7[39];   // BLUNGER TRANSFER DESTINATION
   YP_BLUNGER_WATER_FILL : ALIAS FOR YP_T21[1];
   YP_C5 : COUNTER[15] := ([10].PRE := 10000);
   YP_COMMS_FROM_FullersFV : MESSAGE;
        MessageParameters(ServiceCode := 16#0fa2, LocalElement := YP_N10[10], ...)
   YP_COMMS_FROM_MVFVCIP : MESSAGE;
        MessageParameters(ServiceCode := 16#004c, LocalElement := YP_N14[0], ...)
   YP_COMMS_READ_TIMER : ALIAS FOR YP_T21[3];
   YP_CONV_STOP : PlantItem;   // CONV_STOP
   YP_CONV_STOP_RawInput : ALIAS FOR RIO_Rack_3:2:I.Data.7;   // YP_CONV_STOP
   YP_CONVEYOR_STOP_PB_FLG : ALIAS FOR YP_B3[1].7;
   YP_COPY_OF_SELEC_TIMER : ALIAS FOR YP_N55[40];
   YP_DRAIN_RUNNING : ALIAS FOR YP_N40[3].1;
   YP_DRAIN_TIMER_1_SP : ALIAS FOR YP_N55[42];   // Blunger Drain Timer 1
   YP_DRAIN_TIMER_2_SP : ALIAS FOR YP_N55[43];   // Blunger Drain Timer 2
   YP_DRAIN_TIMER_3_SP : ALIAS FOR YP_N55[44];   // Blunger Drain Timer 3
   YP_INP1 : PlantItem;   // INP1
   YP_INP10 : PlantItem;   // INP10
   YP_INP10_RawInput : ALIAS FOR RIO_Rack_3:2:I.Data.14;   // YP_INP10
   YP_INP11 : PlantItem;   // INP11
   YP_INP11_RawInput : ALIAS FOR RIO_Rack_3:2:I.Data.15;   // YP_INP11
   YP_INP1_RawInput : ALIAS FOR RIO_Rack_3:2:I.Data.2;   // YP_INP1
   YP_INP2 : PlantItem;   // INP2
   YP_INP2_RawInput : ALIAS FOR RIO_Rack_3:2:I.Data.3;   // YP_INP2
   YP_INP3 : PlantItem;   // INP3
   YP_INP3_RawInput : ALIAS FOR RIO_Rack_3:2:I.Data.4;   // YP_INP3
   YP_INP4 : PlantItem;   // INP4
   YP_INP4_RawInput : ALIAS FOR RIO_Rack_3:2:I.Data.8;   // YP_INP4
   YP_INP5 : PlantItem;   // INP5
   YP_INP5_RawInput : ALIAS FOR RIO_Rack_3:2:I.Data.9;   // YP_INP5
   YP_INP6 : PlantItem;   // INP6
   YP_INP6_RawInput : ALIAS FOR RIO_Rack_3:2:I.Data.10;   // YP_INP6
   YP_INP7 : PlantItem;   // INP7
   YP_INP7_RawInput : ALIAS FOR RIO_Rack_3:2:I.Data.11;   // YP_INP7
   YP_INP8 : PlantItem;   // INP8
   YP_INP8_RawInput : ALIAS FOR RIO_Rack_3:2:I.Data.12;   // YP_INP8
   YP_INP9 : PlantItem;   // INP9
   YP_INP9_RawInput : ALIAS FOR RIO_Rack_3:2:I.Data.13;   // YP_INP9
   YP_N10 : INT[105] := ([0] := 1, [10] := 1);   // COMMS BLOC comms block to fv pl c
   YP_N114 : INT[261];   // Original N File From SLC, No Description Available
   YP_N14 : INT[135] := ([103] := 3011, [113] := 3011);   // Original N File From SLC, No Description Available
        [101].0   // Yeast Press Ch1 CIP Active
        [103]   // Yeast Press Ch1 CIP Fault
        [104].0   // Yeast Press Ch1 CIP Route Open
        [111].0   // Yeast Press Ch2 CIP Active
        [113]   // Yeast Press Ch2 CIP Fault
        [114].0   // Yeast Press Ch1 CIP Route Open
   YP_N32 : INT[257];
   YP_N40 : INT[9] := ([0] := 1, [1] := 1, [2] := 1, [3] := 1);   // Original N File From SLC, No Description Available
        [0].0   // Ready to close
        [0].1   // Press Closing
        [0].4   // Press Feed
        [0].5   // Cycle Ended
        [0].6   // Ready for discharge
        [0].7   // Press Opening
        [0].8   // Conveyor discharge
        [1].0   // Conveyor discharging
        [1].2   // Yeast Press Set for CIP ?
        [1].3   // Yeast Press CIP Pulsing ?
        [1].4   // CIP Complete
        [2].0   // BLUNGER WATER FILL IDLE
        [2].1   // Blunger Water Feed Running
        [3].0   // BLUNGER DRAIN/RANSFER TO YST IDLE FLAG
   YP_N50 : INT[15];   // Original N File From SLC, No Description Available
   YP_N55 : INT[244];   // Original N File From SLC, No Description Available
        [0]   // Status 0=Filtration 1=CIP
        [12]   // CIP Variables CIP Valve Change
        [13]   // CIP Variables CIP Total Cycle Time
        [20]   // Fill Cycle Variables Lower Filtrate Valve
        [21]   // Fill Cycle Variables Feed Cycle Timer
        [22]   // Fill Cycle Variables End of Cycle Pause
        [31]   // BLUNGER FILL TIMER SELECTED FROM PV
        [32]   // Blunger Water Feed Feed Timer 1
        [33]   // Blunger Water Feed Feed Timer 2
        [34]   // Blunger Water Feed Feed Timer 3
        [41]   // Blunger Drain Timer Select
        [42]   // Blunger Drain Timer 1
        [43]   // Blunger Drain Timer 2
        [44]   // Blunger Drain Timer 3
   YP_N7 : INT[56] := ([40] := 3);   // INTEGER
        [39]   // BLUNGER TRANSFER DESTINATION
        [40].0   // YST1 HIGH LEVEL FLAG ON=WET
        [40].1   // YST2 HIGH LEVEL FLAG ON=WET
   YP_N88 : INT[7];   // Original N File From SLC, No Description Available
   YP_NO_TANK_SELECTED : ALIAS FOR YP_N7[38].2;
   YP_OUT1 : PlantItem;   // OUT1
   YP_OUT1_ALARM : ALARM_DIGITAL;
   YP_OUT1_DR : ALIAS FOR RIO_Rack_3:3:O.Data.0;
   YP_OUT2 : PlantItem;   // OUT2
   YP_OUT2_ALARM : ALARM_DIGITAL;
   YP_OUT2_DR : ALIAS FOR RIO_Rack_3:3:O.Data.1;
   YP_OUT3 : PlantItem;   // OUT3
   YP_OUT3_ALARM : ALARM_DIGITAL;
   YP_OUT3_DR : ALIAS FOR RIO_Rack_3:3:O.Data.2;
   YP_OUT4 : PlantItem;   // OUT4
   YP_OUT4_ALARM : ALARM_DIGITAL;
   YP_OUT4_DR : ALIAS FOR RIO_Rack_3:3:O.Data.4;
   YP_OUT5 : PlantItem;   // OUT5
   YP_OUT5_ALARM : ALARM_DIGITAL;
   YP_OUT5_DR : ALIAS FOR RIO_Rack_3:3:O.Data.12;
   YP_OUT6 : PlantItem;   // OUT6
   YP_OUT6_ALARM : ALARM_DIGITAL;
   YP_OUT6_DR : ALIAS FOR RIO_Rack_3:3:O.Data.13;
   YP_OUT7 : PlantItem;   // OUT7
   YP_OUT7_ALARM : ALARM_DIGITAL;
   YP_OUT7_DR : ALIAS FOR RIO_Rack_3:3:O.Data.15;
   YP_PILZ_OK : PlantItem;   // PILZ_OK
   YP_PILZ_OK_FLAG : ALIAS FOR YP_B3[1].0;
   YP_PILZ_OK_RawInput : ALIAS FOR RIO_Rack_3:2:I.Data.0;   // YP_PILZ_OK
   YP_PRESS_CL : PlantItem;   // PRESS_CL
   YP_PRESS_CL_RawInput : ALIAS FOR RIO_Rack_3:2:I.Data.5;   // YP_PRESS_CL
   YP_PRESS_CLOSE_PB_FLAG : ALIAS FOR YP_B3[1].5;
   YP_PRESS_OP : PlantItem;   // PRESS_OP
   YP_PRESS_OP_RawInput : ALIAS FOR RIO_Rack_3:2:I.Data.6;   // YP_PRESS_OP
   YP_PRESS_OPEN_PB_FLAG : ALIAS FOR YP_B3[1].6;
   YP_SELECTED_FILL_TIMER : ALIAS FOR YP_N55[30];
   YP_START_DRAIN_FROM_PV : ALIAS FOR YP_B103[3].2;
   YP_START_WATER_FILL : ALIAS FOR YP_B103[3].0;   // START BLUNGER WATER FILL FROM PV
   YP_STOP_DRAIN_B_FROM_PV : ALIAS FOR YP_B103[3].3;
   YP_STOP_WATER_FILL : ALIAS FOR YP_B103[3].1;   // STOP BLUNGER WATER FILL FROM PV
   YP_SYSTEM_4_BIT6_TIMEBASE : ALIAS FOR One_Second_1_scan;
   YP_T20 : TIMER[55] := ([0].PRE := 10000, [1].PRE := 10000, [2].PRE := 10000, [3].PRE := 10000, [4].PRE := 10000, [5].PRE := 10000, [6].PRE := 10000, [7].PRE := 10000, [8].PRE := 10000, [9].PRE := 10000, [10].PRE := 10000, [11].PRE := 10000, [12].PRE := 10000, [13].PRE := 10000, [14].PRE := 10000, [15].PRE := 10000, [16].PRE := 60000, [17].PRE := 10000, [18].PRE := 10000, [18].ACC := 10000, [18].EN := 1, [18].DN := 1);